// TIA Portal project "N16-1166-5_27082020" (V13) (continued)

               #IFM_Switch_State := #IFM_Switch_State + 1;
           1:
               // set number of pulses to send to the IFM senzor
               #IFM_Pulse_Number := #IFM_ApplicationIndex;
               //change the state to the next value
               #IFM_Switch_State := #IFM_Switch_State + 1;
           2:
               //pulsing in precisely time intervals
               IF #IFM_Pulse_Number > 0 THEN
                   IF #IFM_Input_2 = false AND #IFM_Timer_State = 0 THEN
                       #IFM_Input_2 := true;
                       #IFM_Timer_State := #IFM_Pulse_Period / 2;
                   ELSIF #IFM_Input_2 = true AND #IFM_Timer_State = 0 THEN
                       #IFM_Input_2 := false;
                       #IFM_Timer_State := #IFM_Pulse_Period / 2;
                       #IFM_Pulse_Number := #IFM_Pulse_Number - 1;
                   END_IF;
               ELSE
                   #IFM_Switch_State := #IFM_Switch_State + 1;
               END_IF;
           3:
               // set input 1 to false
               #IFM_Input_1 := false;
               //set to init state
               #IFM_Switch_State := 0;
               //set free to switch of application       
               #IFM_PulsApplicationSwitch := true;
           ELSE  // Statement section ELSE
               #IFM_Switch_State := 0;
               #IFM_Input_1 := false;
               #IFM_Input_2 := false;
       END_CASE;
   ELSE
       #IFM_PulsApplicationSwitch := false;
   END_IF;
   *)
END_FUNCTION_BLOCK

FUNCTION_BLOCK "vacuum_cleaner_controll"   // FB2, SCL
{ S7_Optimized_Access := 'FALSE' }
VERSION : 0.1
BEGIN

   IF #vacuum_sensor = true THEN
       #switch := true;
       #timer_lib_Instance.lock := false;
       #vacuum_control_variable := true;
   END_IF;

   IF #switch = true THEN
       #timer_lib_Instance(time_value := #vacuum_cleaner_activity_interval);
       IF #timer_lib_Instance.DONE = true THEN
           #switch := false;
           #vacuum_control_variable := false;
       END_IF;
   END_IF;
END_FUNCTION_BLOCK

FUNCTION_BLOCK "RPA30_F_TRIGR"   // FB4, SCL
{ S7_Optimized_Access := 'FALSE' }
VERSION : 0.1
BEGIN

   IF #PREVIOS = true AND #CLK = false THEN
       #Q := true;
       #STATE := true;
   ELSE
       #Q := false;
   END_IF;

   #PREVIOS := #CLK;
END_FUNCTION_BLOCK

FUNCTION_BLOCK "PA30_IFM_point_checking"   // FB5, SCL
{ S7_Optimized_Access := 'FALSE' }
VERSION : 0.1
BEGIN




   IF #execute = true THEN
   (*
   ** if keyence are disabled in its checking
   *)
       IF #checking_state >= 30 AND #keyence_enable = false THEN
           #checking_state := 27;
       END_IF;

       #index := 0;
       #mark := 0;
       #temp_string := '';

       //pars input data from left ifm sensor 
       WHILE #index < "RPA30_DataBlock".pa30_right_size_in DO
           IF "RPA30_DataBlock".pa30_left_ifm_data[#index] = '#' THEN
               IF #mark > 1 THEN
                   #left_camera_points_pixel[#mark - 1] := STRING_TO_UINT(#temp_string);
                   #temp_string := '';
               END_IF;

               #mark := #mark + 1;
           ELSE
               IF #mark > 1 THEN
                   #temp_string := CONCAT(IN1 := #temp_string, IN2 := "RPA30_DataBlock".pa30_left_ifm_data[#index]);
               END_IF;
           END_IF;

           #index := #index + 1;
       END_WHILE;

       #index := 0;
       #mark := 0;
       #temp_string := '';

       //pars input data from right ifm sensor
       WHILE #index < "RPA30_DataBlock".pa30_right_size_in DO
           IF "RPA30_DataBlock".pa30_right_ifm_data[#index] = '#' THEN
               IF #mark > 1 THEN
                   #right_camera_points_pixel[#mark - 1] := STRING_TO_UINT(#temp_string);
                   #temp_string := '';
               END_IF;

               #mark := #mark + 1;
           ELSE
               IF #mark > 1 THEN
                   #temp_string := CONCAT(IN1 := #temp_string, IN2 := "RPA30_DataBlock".pa30_right_ifm_data[#index]);
               END_IF;
           END_IF;

           #index := #index + 1;
       END_WHILE;

       IF #ifm_side > 0 THEN
           CASE #checking_state OF
               0, 1:  // nastavení senzorů
                   #DONE := false;
                   #checking_state := 2;

               2:
   (* kontrola zda byla aplikace přepnuta *)
                   IF 1 = "RPA30_DataBlock".pa30_left_ifm_actived_application_index AND
                       1 = "RPA30_DataBlock".pa30_right_ifm_actived_application_index THEN
                       #checking_state := 3;
                   END_IF;

               3:
   (* čekání na deaktivaci senzoru *)
                   IF #left_camera_points_pixel[((#ifm_side - 1) * 2) + 1] = 0 THEN
                       #checking_state := 4;
                   END_IF;

               4:
   (* čekání na aktivaci senzoru na bodě L1 a následné přepnutí kamery na bod L2*)
                   IF #left_camera_points_pixel[((#ifm_side - 1) * 2) + 1] > #pixel_treshold THEN
                       #checking_state := 5;
                       #beep := true;
                       #points := 1;
                   END_IF;

               5:
   (* čekání na deaktivaci senzoru *)
                   IF (#left_camera_points_pixel[((#ifm_side - 1) * 2) + 1] = #left_camera_points_pixel[((#ifm_side - 1) * 2) + 2]) = 0 THEN
                       #checking_state := 6;
                   END_IF;

               6:
   (* čekání na aktivaci senzoru  *)
                   IF #left_camera_points_pixel[((#ifm_side - 1) * 2) + 2] > #pixel_treshold THEN
                       #checking_state := 7;
                       #beep := true;
                       #points := 2;
                   END_IF;
               7:
   (* čekání na deaktivaci obou senzorů *)
                   IF (#left_camera_points_pixel[((#ifm_side - 1) * 2) + 2] + #right_camera_points_pixel[((#ifm_side - 1) * 3) + 1]) = 0 THEN
                       #checking_state := 8;
                   END_IF;

               8:
   (* čekání na aktivaci obou senzorů a následné přepnutí senzoru na bod P2 *)
                   IF #right_camera_points_pixel[((#ifm_side - 1) * 3) + 1] > #pixel_treshold THEN
                       #beep := true;
                       #points := 3;
                       #checking_state := 9;
                   END_IF;
               9:
                   IF (#right_camera_points_pixel[((#ifm_side - 1) * 3) + 1] + #right_camera_points_pixel[((#ifm_side - 1) * 3) + 2]) = 0 THEN
                       #checking_state := 10;
                   END_IF;
               10:
                   IF #right_camera_points_pixel[((#ifm_side - 1) * 3) + 2] > #pixel_treshold THEN
                       #beep := true;
                       #points := 4;
                       #checking_state := 11;
                   END_IF;

               11:
                   IF (#right_camera_points_pixel[((#ifm_side - 1) * 3) + 2] + #right_camera_points_pixel[((#ifm_side - 1) * 3) + 3]) = 0 THEN
                       #checking_state := 12;
                   END_IF;
               12:
                   IF #right_camera_points_pixel[((#ifm_side - 1) * 3) + 3] > #pixel_treshold THEN
                       #beep := true;
                       #points := 5;

                       IF #ifm_side = 2 OR "RPA30_DataBlock".RPA30_station_configuration = 0 THEN
                           #checking_state := 27;
                       ELSE
                           IF #keyence_enable = true THEN
                               #checking_state := 30;
                           ELSE
                               #checking_state := 27;
                           END_IF;
                       END_IF;
                   END_IF;
               30:
                   //sensor 1 non active
                   IF (#ifm_side = 1 AND "RPA30_keyence_left_1" = false) OR (#ifm_side = 3 AND "RPA30_keyence_left_2" = false) THEN
                       #checking_state := 31;
                   END_IF;
               31:
                   //sensor 1 active
                   IF (#ifm_side = 1 AND "RPA30_keyence_left_1" = true) OR #ifm_side = 3 AND "RPA30_keyence_left_2" = true THEN
                       #checking_state := 32;
                       #points := 6;
                       #beep := true;
                   END_IF;
               32:
                   //sensor 1 non active
                   IF (#ifm_side = 1 AND "RPA30_keyence_left_1" = false) OR (#ifm_side = 3 AND "RPA30_keyence_left_2" = false) THEN
                       #checking_state := 33;
                   END_IF;

               33:
                   //sensor 2 non active
                   IF (#ifm_side = 1 AND "RPA30_keyence_middle_2" = false) OR (#ifm_side = 3 AND "RPA30_keyence_middle_1" = false) THEN
                       #checking_state := 34;
                   END_IF;

               34:
                   //sensor 2 active
                   IF (#ifm_side = 1 AND "RPA30_keyence_middle_2" = true) OR #ifm_side = 3 AND ("RPA30_keyence_middle_1" = true) THEN
                       #checking_state := 35;
                       #points := 7;
                       #beep := true;
                   END_IF;
               35:
                   //sensor 2 non active
                   IF (#ifm_side = 1 AND "RPA30_keyence_middle_2" = false) OR (#ifm_side = 3 AND "RPA30_keyence_middle_1" = false) THEN
                       #checking_state := 36;
                   END_IF;
               36:
                   //sensor 3 non active
                   IF (#ifm_side = 1 AND "RPA30_keyence_right_1" = false) OR (#ifm_side = 3 AND "RPA30_keyence_right_2" = false) THEN
                       #checking_state := 37;
                   END_IF;
               37:
                   //sensor 3 atvite
                   IF (#ifm_side = 1 AND "RPA30_keyence_right_1" = true) OR (#ifm_side = 3 AND "RPA30_keyence_right_2" = true) THEN
                       #checking_state := 27;
                       #points := 8;
                       #beep := true;
                   END_IF;
               27:
                   #DONE := true;
          END_CASE;
      END_IF;
   ELSE
       #checking_state := 0;
       #points := 0;
       #DONE := false;
   END_IF;

   (* pípnutí při zachycení bodu *)
   IF #beep = true THEN
       #timer_lib_Instance(100);
       IF #timer_lib_Instance.DONE = false THEN
           #primerbox_siren := true;
       ELSE
           #primerbox_siren := false;
           #beep := false;
       END_IF;
   END_IF;
END_FUNCTION_BLOCK

FUNCTION_BLOCK "O2VxEth1500"   // FB8, SCL
TITLE = O2VxEth1500 for S7-15xx CPU FW V1.7 or higher
{ S7_Optimized_Access := 'FALSE' }
AUTHOR : ifm-sytl
FAMILY : O2Vx
NAME : O2Vx1500
VERSION : 1.3
// Basic Application program for O2Vx
// connected to S7-1500 station via CPU-internal Ethernet interface
// for S7-15xx CPU Firmware V1.7 or higher
BEGIN
END_FUNCTION_BLOCK

FUNCTION_BLOCK "fs_scaner_fce"   // FB11, SCL
{ S7_Optimized_Access := 'FALSE' }
VERSION : 0.1
BEGIN
   #Receive_P2P_Instance(BUFFER:=#Receive_P2P_Instance.ReceiveBuffer,"PORT" := "FS~CM_PtP_1");

   IF #Receive_P2P_Instance.NDR = true THEN
      Chars_TO_Strg(Chars:=#Receive_P2P_Instance.ReceiveBuffer,
                    pChars:=0,
                    Cnt:=#Receive_P2P_Instance.received_length-1,
                    Strg=>#scaner_input_data);
   END_IF;
END_FUNCTION_BLOCK

FUNCTION_BLOCK "print_label_PA60"   // FB13, SCL
{ S7_Optimized_Access := 'FALSE' }
VERSION : 0.1
BEGIN

   #DONE := false;

   IF #TCON_Instance.DONE = false THEN
       #TCON_Instance.REQ := NOT #TCON_Instance.REQ;
       #TCON_Instance(CONNECT := "printer_connection",
                               ID := 10);
   ELSE
       //date formating
       #date_string := CONCAT(IN1 := #date_string, IN2 := "copyAndFill"(characterFill := '0', charReplace := '+', stringIn := (DELETE(IN := INT_TO_STRING(#"date".DAY), L := 1, P := 1)), P := 0, char_number := 2));
       #date_string := CONCAT(IN1 := #date_string, IN2 := '.');
       #date_string := CONCAT(IN1 := #date_string, IN2 := "copyAndFill"(characterFill := '0', charReplace := '+', stringIn := (DELETE(IN := INT_TO_STRING(#"date".MONTH), L := 1, P := 1)), P := 0, char_number := 2));
       #date_string := CONCAT(IN1 := #date_string, IN2 := '.');
       #date_string := CONCAT(IN1 := #date_string, IN2 := "copyAndFill"(characterFill := '0', charReplace := '+', stringIn := (DELETE(IN := UINT_TO_STRING(#"date".YEAR), L := 1, P := 1)), P := 0, char_number := 4));

       //time formating
       #time_string := CONCAT(IN1 := #time_string, IN2 := "copyAndFill"(characterFill := '0', charReplace := '+', stringIn := (DELETE(IN := INT_TO_STRING(#"date".HOUR), L := 1, P := 1)), P := 0, char_number := 2));
       #time_string := CONCAT(IN1 := #time_string, IN2 := ':');
       #time_string := CONCAT(IN1 := #time_string, IN2 := "copyAndFill"(characterFill := '0', charReplace := '+', stringIn := (DELETE(IN := INT_TO_STRING(#"date".MINUTE), L := 1, P := 1)), P := 0, char_number := 2));
       #time_string := CONCAT(IN1 := #time_string, IN2 := ':');
       #time_string := CONCAT(IN1 := #time_string, IN2 := "copyAndFill"(characterFill := '0', charReplace := '+', stringIn := (DELETE(IN := INT_TO_STRING(#"date".SECOND), L := 1, P := 1)), P := 0, char_number := 2));

       //qr code string formating
       IF #frame_conf = 0 THEN
           #MCode := 'AU581*1762975*';
       ELSE
           #MCode := 'AU326-1*1768362*';
       END_IF;

       #MCode := CONCAT(IN1 := #MCode, IN2 := #date_string);
       #MCode := CONCAT(IN1 := #MCode, IN2 := '*');
       #MCode := CONCAT(IN1 := #MCode, IN2 := #time_string);
       #MCode := CONCAT(IN1 := #MCode, IN2 := '*172');
       #MCode := CONCAT(IN1 := #MCode, IN2 := #order);

       //send command to the printer
       IF #TSEND_Instance.DONE = false THEN

       #numberOfChar := 0;
       Strg_TO_Chars(Strg := '^XA^MMT^PW480^LL0200^LS0^FO0,0^GFA,03072,03072,00032,:Z64:eJztk7GO4jAQhifJIZ2gIYWbrbZchTdI5Ui3PUjx+1jQ8RRZaCK7uTI3vNz9M4YEpIu47nQSI+wYO1/GM/MP0cte9k/NbXW2c+ehm+Y/8nb8StaOu5m7raKSG5mLMJ3Hv+WT56rHlE88jcvEm1mevcz1IP554nl88QkflF/O+X/GZ1H5VU8V4s/TZh7G+K8v',
                     pChars := #chars,
                     Cnt => #chars,
                     Chars := #data_out);

       #numberOfChar := #numberOfChar +#chars;
       Strg_TO_Chars(Strg := 'mi0+lLXGUoYvGSfb7sF/HvALPS1D8CEc5V9/zy9cmznXknPGOvfp2kWqbIr/bXhjzi/MVDN75iMPWFz5THjj4NQ58K5RHhvJPzzCfxXCPqhvecI/Nrzy39S/s8Kl0RJ4pzzix4vdqo9+c4jneIgxHgIV8R0L5W1ZlmvwZBp4b3CLzxbbGZaSWvUalj3ucApU7dNA/oOvurv8C9+SAYvLK09GjvgofP2Lmc+IXsaBO7pAATV4eIT/0uxw3V3ic',
                     pChars := #numberOfChar,
                     Cnt => #chars,
                     Chars := #data_out);

       #numberOfChar := #numberOfChar + #chars;
       Strg_TO_Chars(Strg := 'Q+kEsVUPpyEr3pMJ2Qfo/KSBohhqfwPSYB75CWMKx+V33wh3HNPGxk+xq+IZlgpvyspW4NX/ShvzR0vNac+dEH1V0kOfC5/sVA+9W8z8cjIHV8PeOuDOxQ7R8gnDE/1T77Fb0S0Jao35d8S0oH8aWqvneeR7n24agCeVQj+xi/Ap/qLhhqQt/rTSjqlQPWj1t5HfXax32j9adEmFT7qz476085LKoT+EbTewav+5GSR4qeb/o2T/J',
                     pChars := #numberOfChar,
                     Cnt => #chars,
                     Chars := #data_out);

       #numberOfChar := #numberOfChar + #chars;
       Strg_TO_Chars(Strg := 'PoX9sxH7QLEPxQMA9UX1B/aYOC9SRTXhQnjWfxPfTPVsJKysolSYRLVLjtEkt5YHT0PTWwTfysKf8xf678ev5c7f3J+cte9rL/zn4DEoMnnA==:C58E',
                     pChars := #numberOfChar,
                     Cnt => #chars,
                     Chars := #data_out);

       #numberOfChar := #numberOfChar + #chars;
       IF #frame_conf = 0 THEN
           Strg_TO_Chars(Strg := '^FT32,85^A0N,17,16^FH\^FDAU581^FS^FT32,104^A0N,17,16^FH\^FDID-No. 1762975^FS^FT180,122^A0N,17,16^FH\^FD',
                         pChars := #numberOfChar,
                         Cnt => #chars,
                         Chars := #data_out);
       ELSE //zde upravit kód rámu
           Strg_TO_Chars(Strg := '^FT32,85^A0N,17,16^FH\^FDAU326-1^FS^FT32,104^A0N,17,16^FH\^FDID-No. 1768362^FS^FT180,122^A0N,17,16^FH\^FD',
                         pChars := #numberOfChar,
                         Cnt => #chars,
                         Chars := #data_out);
       END_IF;

       #numberOfChar := #numberOfChar + #chars;
       Strg_TO_Chars(Strg := #time_string,
                     pChars := #numberOfChar,
                     Cnt => #chars,
                     Chars := #data_out);

       #numberOfChar := #numberOfChar + #chars;
       Strg_TO_Chars(Strg := '^FS^FT31,142^A0N,17,16^FH\^FDSerial-No:^FS',
                         pChars := #numberOfChar,
                         Cnt => #chars,
                         Chars := #data_out);

       #numberOfChar := #numberOfChar + #chars;
       Strg_TO_Chars(Strg := '^BY96,96^FT332,141^BXN,4,200,0,0,1,~^FH\^FD',
                     pChars := #numberOfChar,
                     Cnt => #chars,
                     Chars := #data_out);

       #numberOfChar := #numberOfChar + #chars;
       Strg_TO_Chars(Strg := #MCode,
                     pChars := #numberOfChar,
                     Cnt => #chars,
                     Chars := #data_out);

       #numberOfChar := #numberOfChar + #chars;
       Strg_TO_Chars(Strg := '^FS^FT32,161^A0N,17,16^FH\^FDWBR Made in Romania (WRO)^FS^FT31,123^A0N,17,16^FH\^FDDate:^FS^FT31,181^A0N,17,16^FH\^FD',
                     pChars := #numberOfChar,
                     Cnt => #chars,
                     Chars := #data_out);

       #numberOfChar := #numberOfChar + #chars;
       Strg_TO_Chars(Strg := #MCode,
                     pChars := #numberOfChar,
                     Cnt => #chars,
                     Chars := #data_out);

       #numberOfChar := #numberOfChar + #chars;
       Strg_TO_Chars(Strg := '^FS^FT70,122^A0N,17,16^FH\^FD',
                     pChars := #numberOfChar,
                     Cnt => #chars,
                     Chars := #data_out);

       #numberOfChar := #numberOfChar + #chars;
       Strg_TO_Chars(Strg := #date_string,
                     pChars := #numberOfChar,
                     Cnt => #chars,
                     Chars := #data_out);

       #numberOfChar := #numberOfChar + #chars;
       Strg_TO_Chars(Strg := '^FS^FT179,142^A0N,17,16^FH\^FD',
                     pChars := #numberOfChar,
                     Cnt => #chars,
                     Chars := #data_out);

       #numberOfChar := #numberOfChar + #chars;
       Strg_TO_Chars(Strg := #order,
                     pChars := #numberOfChar,
                     Cnt => #chars,
                     Chars := #data_out);

       #numberOfChar := #numberOfChar + #chars;
       Strg_TO_Chars(Strg := '^FS^FT114,142^A0N,17,16^FH\^FD172^FS^PQ1,0,1,Y^XZ',
                     pChars := #numberOfChar,
                     Cnt => #chars,
                     Chars := #data_out);

       #numberOfChar := #numberOfChar + #chars;


           #TSEND_Instance.REQ := NOT #TSEND_Instance.REQ;
           #TSEND_Instance(ID := 10,LEN := #numberOfChar, DATA := #data_out);
       ELSE
           IF #TDISCON_Instance.DONE = false THEN
               #TDISCON_Instance.REQ := NOT #TDISCON_Instance.REQ;
               #TDISCON_Instance(ID := 10);
           ELSE
               #TDISCON_Instance.DONE := false;
               #TSEND_Instance.DONE := false;
               #TCON_Instance.DONE := false;
               #DONE := true;
           END_IF;
       END_IF;
   END_IF;
END_FUNCTION_BLOCK

FUNCTION_BLOCK "bottle_changing"   // FB14, SCL
{ S7_Optimized_Access := 'FALSE' }
VERSION : 0.1
BEGIN

   #DONE := false;

   CASE #"step" OF
      0:  // take secound bottle than will used
          IF #bottle = 1 THEN
              #hmi_label_index := 28;
              #use_bottle_2 := true ;
              #use_bottle_1 := false;
          ELSIF #bottle = 2 THEN
              #hmi_label_index := 29;
              #use_bottle_2 := false;
              #use_bottle_1 := true;
          END_IF;



          IF (#bottle_presence_sensor_1 = false AND  #bottle = 2) OR (#bottle_presence_sensor_2 = false AND  #bottle = 1) THEN
              #"step" := 10;
              #take_bottle := true;
          END_IF;

      10: // scan label and check expiration
          #hmi_label_index := "RPA10B_hmi_scan_bottle";
          IF "RPA10B_Scanner_DB".NDR = true THEN
              IF RD_SYS_T(#current_time) < 0 THEN
                  ;
              END_IF;

              #bottle_checking_result := "bottle_label_check"(input_data := "RPA10B_datablock".RPA10B_scanned_data, chemical_type := 5);

              IF #bottle_checking_result = 0 THEN
                  IF  #bottle_presence_sensor_2 = false  THEN
                      #bottle_label_2 := "RPA10B_datablock".RPA10B_scanned_data;
                  ELSIF #bottle_presence_sensor_1 = false THEN
                      #bottle_label_1 := "RPA10B_datablock".RPA10B_scanned_data;
                  END_IF;

                  IF (#bottle = 1 AND #bottle_presence_sensor_2 = false) OR (#bottle = 2 AND #bottle_presence_sensor_2 = false) THEN
                      #"step" := 40;
                  ELSIF (#bottle = 1 AND #bottle_presence_sensor_1 = false) OR (#bottle = 2 AND #bottle_presence_sensor_1 = false) THEN
                      #"step" := 20;
                  END_IF;

              ELSIF #bottle_checking_result = 2 THEN
                  "RPA10B_datablock".PA10B_error_state_lock := 400;
                  #"step" := 30;
              ELSIF #bottle_checking_result = 3 THEN
                  "RPA10B_datablock".PA10B_error_state_lock := 401;
                  #"step" := 30;
              ELSIF #bottle_checking_result = 4 THEN
                  "RPA10B_datablock".PA10B_error_state_lock := 402;
                  #"step" := 30;
              ELSIF #bottle_checking_result = 5 THEN
                  "RPA10B_datablock".PA10B_error_state_lock := 403;
                  #"step" := 30;
              END_IF;
          END_IF;

      20: //change pad bottle 1
          #hmi_label_index := "RPA10B_hmi_change_pad";
          "RPA10B_datablock".RPA10B_show_pad_left := true;
          IF "RPA10B_change_pad"(padSensor := "RPA10B_primerbox_pad_sensor_left",
                                     padIsChangedButton := "RPA10B_primerbox_button_PAD_IS_CHANGED",
                                     failStatelockIdetifier := 6,
                                     bigFailStateLock := "RPA10B_datablock".PA10B_big_fail_state_lock,
                                     FatalErrorStateLock := "RPA10B_datablock".PA10B_fatal_error_state_lock,
                                     readyLED => "RPA10B_primerbox_LED_green_ready",
                                     notReadyLED => "RPA10B_primerbox_LED_red_NOT_READY",
                                     changePedLED => "RPA10B_primerbox_LED_orange_change_pad",
                                     confirmButtonLED => "RPA10B_LCD_LED_blue_confirm_button",
                                     failStateLock := "RPA10B_datablock".PA10B_fail_state_lock) THEN
              "RPA10B_datablock".RPA10B_show_pad_left := false;
              #bottle_1_cyclus_counter := 0;
              IF RD_SYS_T(#bottle_1_expiration) < 2 THEN
                  IF (#bottle = 2 AND #bottle_presence_sensor_1 = false) OR (#bottle = 1 AND #bottle_presence_sensor_2 = false) THEN
                      #"step" := 50;
                  ELSE
                      #"step" := 60;
                  END_IF;
              END_IF;
          END_IF;

      30: // bottle expired
          IF "RPA10B_datablock".PA10B_error_state_lock = 400 OR "RPA10B_datablock".PA10B_error_state_lock = 401 OR "RPA10B_datablock".PA10B_error_state_lock = 402 OR "RPA10B_datablock".PA10B_error_state_lock = 403 THEN
              "RPA10B_LCD_LED_blue_confirm_button" := "Clock_0.5Hz";
              IF "RPA10B_LCD_button_confirm" = true THEN
                  "RPA10B_datablock".PA10B_error_state_lock := 0;
                  "RPA10B_LCD_LED_blue_confirm_button" := false;
                  #"step" := 10;
              END_IF;
          END_IF;

      40: // change pad bottle 2
          #hmi_label_index := "RPA10B_hmi_change_pad";
          "RPA10B_datablock".RPA10B_show_pad_right := true;
          IF "RPA10B_change_pad"(padSensor := "RPA10B_primerbox_pad_sensor_right",
                                     padIsChangedButton := "RPA10B_primerbox_button_PAD_IS_CHANGED",
                                     failStatelockIdetifier := 6,
                                     bigFailStateLock := "RPA10B_datablock".PA10B_big_fail_state_lock,
                                     FatalErrorStateLock := "RPA10B_datablock".PA10B_fatal_error_state_lock,
                                     readyLED => "RPA10B_primerbox_LED_green_ready",
                                     notReadyLED => "RPA10B_primerbox_LED_red_NOT_READY",
                                     changePedLED => "RPA10B_primerbox_LED_orange_change_pad",
                                     confirmButtonLED => "RPA10B_LCD_LED_blue_confirm_button",
                                     failStateLock := "RPA10B_datablock".PA10B_fail_state_lock) THEN
              "RPA10B_datablock".RPA10B_show_pad_right := false;
              #bottle_2_cyclus_counter := 0;
              IF RD_SYS_T(#bottle_2_expiration) < 2 THEN
                  IF (#bottle = 1 AND #bottle_presence_sensor_2 = false) OR (#bottle = 2 AND #bottle_presence_sensor_1 = false) THEN
                      #"step" := 50;
                  ELSE
                      #"step" := 60;
                  END_IF;
              END_IF;
          END_IF;

      50: // put bottle back to primerbox and take secound bottle
          IF #bottle_presence_sensor_1 = true AND #bottle_presence_sensor_2 = true THEN
              #take_bottle := false;
              IF #bottle = 1 THEN
                  //choose bottle 1
                  #hmi_label_index := 28;
                  #use_bottle_2 := false;
                  #use_bottle_1 := true;
              ELSIF #bottle = 2 THEN
                  //choose bottle 2
                  #hmi_label_index := 29;
                  #use_bottle_2 := true;
                  #use_bottle_1 := false;
              END_IF;
          ELSE
              //put bottle back to primer box
              #hmi_label_index := 30;
          END_IF;

          IF (#bottle = 1 AND #bottle_presence_sensor_1 = false) OR (#bottle = 2 AND #bottle_presence_sensor_2 = false) THEN
              #take_bottle := true;
              #"step" := 10;
          END_IF;

      60: //end
          #DONE := true;
          #"step" := 0;
       ELSE  // Statement section ELSE
           #"step" := 0;
   END_CASE;
END_FUNCTION_BLOCK

FUNCTION_BLOCK "fs_print_label_fce"   // FB15, SCL
{ S7_Optimized_Access := 'FALSE' }
VERSION : 0.1
BEGIN
END_FUNCTION_BLOCK

FUNCTION_BLOCK "shaker_door_lock_control"   // FB18, SCL
{ S7_Optimized_Access := 'FALSE' }
VERSION : 0.1
BEGIN


   #mixer_1_door_1_lock := #mixer_1_presence_sensor_1 AND #mixer_1_door_1_is_close AND #mixer_door_lock_enable[0];
   #mixer_1_door_2_lock := #mixer_1_presence_sensor_2 AND #mixer_1_door_2_is_close AND #mixer_door_lock_enable[1];
   #mixer_2_door_1_lock := #mixer_2_presence_sensor_1 AND #mixer_2_door_1_is_close AND #mixer_door_lock_enable[2];
   #mixer_2_door_2_lock := #mixer_2_presence_sensor_2 AND #mixer_2_door_2_is_close AND #mixer_door_lock_enable[3];
   #mixer_3_door_1_lock := (#mixer_3_presence_sensor_1 AND #mixer_3_door_1_is_close AND #mixer_door_lock_enable[4]);
END_FUNCTION_BLOCK

FUNCTION_BLOCK "print_label_582"   // FB19, SCL
{ S7_Optimized_Access := 'FALSE' }
VERSION : 0.1
BEGIN





   #DONE := false;

   IF #TCON_Instance.DONE = false THEN
       #TCON_Instance.REQ := NOT #TCON_Instance.REQ;
       #TCON_Instance(CONNECT := "printer_connection",
                               ID := 10);
   ELSE

       //date formating
       #date_string := CONCAT(IN1 := #date_string, IN2 := "copyAndFill"(characterFill := '0', charReplace := '+', stringIn := (DELETE(IN := INT_TO_STRING(#"date".DAY), L := 1, P := 1)), P := 0, char_number := 2));
       #date_string := CONCAT(IN1 := #date_string, IN2 := '.');
       #date_string := CONCAT(IN1 := #date_string, IN2 := "copyAndFill"(characterFill := '0', charReplace := '+', stringIn := (DELETE(IN := INT_TO_STRING(#"date".MONTH), L := 1, P := 1)), P := 0, char_number := 2));
       #date_string := CONCAT(IN1 := #date_string, IN2 := '.');
       #date_string := CONCAT(IN1 := #date_string, IN2 := "copyAndFill"(characterFill := '0', charReplace := '+', stringIn := (DELETE(IN := UINT_TO_STRING(#"date".YEAR), L := 1, P := 1)), P := 0, char_number := 4));

       //time formating
       #time_string := CONCAT(IN1 := #time_string, IN2 := "copyAndFill"(characterFill := '0', charReplace := '+', stringIn := (DELETE(IN := INT_TO_STRING(#"date".HOUR), L := 1, P := 1)), P := 0, char_number := 2));
       #time_string := CONCAT(IN1 := #time_string, IN2 := ':');
       #time_string := CONCAT(IN1 := #time_string, IN2 := "copyAndFill"(characterFill := '0', charReplace := '+', stringIn := (DELETE(IN := INT_TO_STRING(#"date".MINUTE), L := 1, P := 1)), P := 0, char_number := 2));
       #time_string := CONCAT(IN1 := #time_string, IN2 := ':');
       #time_string := CONCAT(IN1 := #time_string, IN2 := "copyAndFill"(characterFill := '0', charReplace := '+', stringIn := (DELETE(IN := INT_TO_STRING(#"date".SECOND), L := 1, P := 1)), P := 0, char_number := 2));

       //qr code string formating
       #MCode := 'AU582*1762976*';
       #MCode := CONCAT(IN1 := #MCode, IN2 := #date_string);
       #MCode := CONCAT(IN1 := #MCode, IN2 := '*');
       #MCode := CONCAT(IN1 := #MCode, IN2 := #time_string);
       #MCode := CONCAT(IN1 := #MCode, IN2 := '*172');
       #MCode := CONCAT(IN1 := #MCode, IN2 := #order_string);

       //command formating
       #command := CONCAT(IN1 := #command, IN2 := '^XA');
       #command := CONCAT(IN1 := #command, IN2 := #label1);
       //...next data in the label

       //barcode
       #command := CONCAT(IN1 := #command, IN2 := '^BY96,96^FT270,145^BXN,4,200,0,0,1,~^FH\^FD');
       #command := CONCAT(IN1 := #command, IN2 := #MCode);
       #command := CONCAT(IN1 := #command, IN2 := '^FS');

       //label
       #command := CONCAT(IN1 := #command, IN2 := '^FT31,181^A0N,16,14^FH\^FD');
       #command := CONCAT(IN1 := #command, IN2 := #MCode);
       #command := CONCAT(IN1 := #command, IN2 := '^FS');

       //date
       #command := CONCAT(IN1 := #command, IN2 := '^FT70,122^A0N,17,16^FH\^FD');
       #command := CONCAT(IN1 := #command, IN2 := #date_string);
       #command := CONCAT(IN1 := #command, IN2 := '^FS');
       Strg_TO_Chars(Strg := #command,
                     pChars := 0,
                     Cnt => #chars,
                     Chars := #data_out);

       #command := '';
       //time
       #command := CONCAT(IN1 := #command, IN2 := '^FT180,122^A0N,17,16^FH\^FD');
       #command := CONCAT(IN1 := #command, IN2 := #time_string);
       #command := CONCAT(IN1 := #command, IN2 := '^FS');

       //order part 1
       #command := CONCAT(IN1 := #command, IN2 := '^FT114,142^A0N,17,16^FH\^FD172^FS');

       //#order part 2
       #command := CONCAT(IN1 := #command, IN2 := '^FT179,142^A0N,17,16^FH\^FD');
       #command := CONCAT(IN1 := #command, IN2 := #order_string);
       #command := CONCAT(IN1 := #command, IN2 := '^FS');

       #command := CONCAT(IN1 := #command, IN2 := '^XZ');

       //prepeare to send

       #numberOfChar := #chars;
       Strg_TO_Chars(Strg := #command,
                     pChars := #chars,
                     Cnt => #chars,
                     Chars := #data_out);

       #numberOfChar := #numberOfChar + #chars;

       //send command to the printer
       IF #TSEND_Instance.DONE = false THEN
           #TSEND_Instance.REQ := NOT #TSEND_Instance.REQ;
           #TSEND_Instance(ID := 1,LEN := #numberOfChar, DATA := #data_out);
       ELSE
           IF #TDISCON_Instance.DONE = false THEN
               #TDISCON_Instance.REQ := NOT #TDISCON_Instance.REQ;
               #TDISCON_Instance(ID := 1);
           ELSE
               #TDISCON_Instance.DONE := false;
               #TSEND_Instance.DONE := false;
               #TCON_Instance.DONE := false;
               #DONE := true;
           END_IF;
       END_IF;
   END_IF;
END_FUNCTION_BLOCK

FUNCTION_BLOCK "scaner_runtime"   // FB20, SCL
{ S7_Optimized_Access := 'FALSE' }
VERSION : 0.1
BEGIN
   #fs_scaner_fce_Instance();


   IF #fs_scaner_fce_Instance.Receive_P2P_Instance.NDR = true THEN
       IF #shaker_index = 0 THEN
           IF #filling_e = false AND #print_sp_bottle_e = false AND #chemical_type > 0 THEN
               IF #fs_scaner_fce_Instance.scaner_input_data[LEN(#fs_scaner_fce_Instance.scaner_input_data)] = 'M' THEN
                   #filling_e := true;
               ELSE
                   #print_sp_bottle_e := true;
               END_IF;
           END_IF;
       END_IF;
   END_IF;
END_FUNCTION_BLOCK

FUNCTION_BLOCK "timer_lib"   // FB21, SCL
{ S7_Optimized_Access := 'FALSE' }
VERSION : 0.1
BEGIN
   #DONE := false;
   IF #lock = true THEN
       IF RD_LOC_T(#actual_time) < 2 THEN
           IF TIME_TO_DINT(IN := T_DIFF(IN1 := #actual_time, IN2 := #"time")) > #time_value THEN
               #DONE := true;
               #lock := false;
           END_IF;
       END_IF;
   ELSE
       IF RD_LOC_T(#"time") < 2 THEN
           #lock := true;
       END_IF;
   END_IF;
END_FUNCTION_BLOCK

FUNCTION_BLOCK "filling_station_main"   // FB23, SCL
{ S7_Optimized_Access := 'FALSE' }
VERSION : 0.1
BEGIN

   IF #fs_activity_state = true THEN
       (* station internal state runtime control *)
       "fs_internal_state"(switch_automat_manual := "ib_FS_LCD_switch_automat_manual",
                           tcp_connection := "tcp_datablock".tcp_connection,
                           confirm_button := "ib_FS_LCD_button_confirm",
                           error_state := #fs_error_state,
                           confirm_led := "ob_FS_LCD_confirm_button_LED_blue",
                           beacon_green := "ob_FS_LCD_beacon_green",
                           beacon_orange := "ob_FS_LCD_beacon_orange",
                           beacon_red := "ob_FS_LCD_beacon_red",
                           beacon_siren := "ob_FS_LCD_beacon_siren",
                           alarm:=#fs_alarm);

       IF #fs_reset_enable = true THEN
           "station_reset"(funel_1:="ob_FS_move_UP_funel_1",
                           funel_2:="ob_FS_move_UP_funel_2",
                           funel_3:="ob_FS_move_UP_funel_3",
                           funel_4:="ob_FS_move_UP_funel_4",
                           funel_5:="ob_FS_move_UP_funel_5",
                           fs_reset_e:=#fs_reset_enable,
                           fs_chemical_type:=#chemical_type,
                           fill_bottle_step:=#fce_filling_Instance."step",
                           shake_deinit:=#sp_bottle_shaking_Instance.shake_deinit,
                           print_sp_bottle_label_step:=#fce_print_sp_botle_label_Instance."step",
                           fs_show_manual_or_scan:=#manual_or_scan,
                           fs_show_button:=#fs_show_button,
                           fs_show_fill_button:=#fce_filling_Instance.show_fill_button,
                           fs_funel_control:=#fce_filling_Instance.funel_control,
                           hmi_label_index:=#hmi_label_index);
       END_IF;

       IF #filling_enable = false AND #print_sp_bottle_label_enable = false AND #shaking_enable = false THEN
           IF #chemical_type > 0 AND #chemical_type < 3 THEN
               #hmi_label_index := 21;
               #fs_show_button := true;
               #manual_or_scan := false;
           ELSIF #chemical_type > 2 THEN
               IF #chemical_type_pre = 0 AND #chemical_type > 2 THEN
                   #manual_or_scan := true;
               END_IF;

               IF #manual_or_scan = false THEN
                   #hmi_label_index := 22;
               ELSE
                   #hmi_label_index := 20;
               END_IF;

               #fs_show_button := true;
           ELSIF #chemical_type = 0 THEN
               #fs_show_button := false;
               #manual_or_scan := false;
               #hmi_label_index := 0;
           END_IF;
       ELSE
           #fs_show_button := true;
           #manual_or_scan := false;
       END_IF;

       #chemical_type_pre := #chemical_type;

       (* scanner runtime hadler and input data parsing *)
       #scaner_runtime_Instance(shaker_index:=#sp_bottle_shaking_Instance.runtime_shaker_index_finding_Instance.shaker_index,
                                chemical_type:=#chemical_type,
                                filling_e:=#filling_enable,
                                print_sp_bottle_e:=#print_sp_bottle_label_enable);

       (* print suplier bottle label work cycle *)
       IF #shaking_enable = false THEN // shaking work cycle is more important
           #fce_print_sp_botle_label_Instance(scanned_data := #scaner_runtime_Instance.fs_scaner_fce_Instance.scaner_input_data,
                                              scaner_ndr := #scaner_runtime_Instance.fs_scaner_fce_Instance.Receive_P2P_Instance.NDR,
                                              expire_time_Primer_DV954V1 := #expire_time_Primer_DV954V1,
                                              expire_time_Activator_DW646 := #expire_time_Activator_DW646,
                                              expire_time_Remover_SIKA_208 := #expire_time_Remover_SIKA_208,
                                              expire_time_Primer_SIKA_207 := #expire_time_Primer_SIKA_207,
                                              expire_time_Activator_SIKA_110 := #expire_time_Activator_SIKA_110,
                                              print_sp_bottle_label_enable := #print_sp_bottle_label_enable,
                                              error_state := #fs_error_state,
                                              fs_SIKA_remover_order := #fs_SIKA_remover_order,
                                              fs_SIKA_primer_order := #fs_SIKA_primer_order,
                                              fs_SIKA_activator_order := #fs_SIKA_activator_order,
                                              shake_enable := #shaking_enable,
                                              chemical_type := #chemical_type,
                                              show_button := #fs_show_button,
                                              hmi_label_index := #hmi_label_index,
                                              show_manual_input := #manual_or_scan);

           (*small bottle filling work cycle*)

           #fce_filling_Instance(scanned_data := #scaner_runtime_Instance.fs_scaner_fce_Instance.scaner_input_data,
                                 scaner_ndr := #scaner_runtime_Instance.fs_scaner_fce_Instance.Receive_P2P_Instance.NDR,
                                 funel_1_bottle_presence := "ib_FS_sensor_bottle_1",
                                 funel_2_bottle_presence := "ib_FS_sensor_bottle_2",
                                 funel_3_bottle_presence := "ib_FS_sensor_bottle_3",
                                 funel_4_bottle_presence := "ib_FS_sensor_bottle_4",
                                 funel_5_bottle_presence := "ib_FS_sensor_bottle_5",
                                 primer_DV954V1_time_after_shaking := #primer_DV954V1_time_after_shaking,
                                 primer_SIKA_207_time_after_shaking := #primer_SIKA_207_time_after_shaking,
                                 filling_enable := #filling_enable,
                                 chemical_type := #chemical_type,
                                 shaking_enable := #shaking_enable,
                                 error_state := #fs_error_state,
                                 move_UP_funel_1 := "ob_FS_move_UP_funel_1",
                                 move_UP_funel_2 := "ob_FS_move_UP_funel_2",
                                 move_UP_funel_3 := "ob_FS_move_UP_funel_3",
                                 move_UP_funel_4 := "ob_FS_move_UP_funel_4",
                                 move_UP_funel_5 := "ob_FS_move_UP_funel_5",
                                 hmi_label_index := #hmi_label_index);

       END_IF;

       (* shaking fce *)


       #sp_bottle_shaking_Instance(shaker_1_door_1_lock := "ob_FS_mixer_1_door_1_lock",
                                   shaker_1_door_2_lock := "ob_FS_mixer_1_door_2_lock",
                                   shaker_2_door_1_lock := "ob_FS_mixer_2_door_1_lock",
                                   shaker_2_door_2_lock := "ob_FS_mixer_2_door_2_lock",
                                   shaker_3_door_1_lock := "ob_FS_mixer_3_door_lock",
                                   chemical_type := #chemical_type,
                                   error_state := #fs_error_state,
                                   shaker_1_door_1_bottle_presence := "ib_FS_mixer_1_presence_sensor_1",
                                   shaker_1_door_2_bottle_presence := "ib_FS_mixer_1_presence_sensor_2",
                                   shaker_2_door_1_bottle_presence := "ib_FS_mixer_2_presence_sensor_1",
                                   shaker_2_door_2_bottle_presence := "ib_FS_mixer_2_presence_sensor_2",
                                   shaker_3_door_1_bottle_presence := "ib_FS_mixer_3_bottle_pressence",
                                   shaker_1_door_1_position := "ib_FS_mixer_1_door_1_is_close",
                                   shaker_1_door_2_position := "ib_FS_mixer_1_door_2_is_close",
                                   shaker_2_door_1_position := "ib_FS_mixer_2_door_1_is_close",
                                   shaker_2_door_2_position := "ib_FS_mixer_2_door_2_is_close",
                                   shaker_3_door_1_position := "ib_FS_mixer_3_door_position",
                                   shaking_enable := #shaking_enable,
                                   scaner_ndr := #scaner_runtime_Instance.fs_scaner_fce_Instance.Receive_P2P_Instance.NDR,
                                   scanned_data := #scaner_runtime_Instance.fs_scaner_fce_Instance.scaner_input_data,
                                   hmi_label_index := #hmi_label_index);


   ELSE
       (* inactive station state *)
       "station_inactive_state"(fs_start_button:="ib_FS_LCD_button_start",
                                fune_1:="ob_FS_move_UP_funel_1",
                                fune_2:="ob_FS_move_UP_funel_2",
                                fune_3:="ob_FS_move_UP_funel_3",
                                fune_4:="ob_FS_move_UP_funel_4",
                                fune_5:="ob_FS_move_UP_funel_5",
                                fs_reset_enable:=#fs_reset_enable,
                                fs_start_led:="ob_FS_LCD_start_button_LED_green",
                                error_state:=#fs_error_state,
                                beacon_red:="ob_FS_LCD_beacon_red",
                                beacon_orange:="ob_FS_LCD_beacon_orange",
                                beacon_green:="ob_FS_LCD_beacon_green",
                                beacon_siren:="ob_FS_LCD_beacon_siren",
                                fs_station_activity:=#fs_activity_state,
                                chemical_type:=#chemical_type,
                                fill_bottle_step:=#fce_filling_Instance."step",
                                shake_deinit:=#sp_bottle_shaking_Instance.shake_deinit,
                                print_sp_bottle_label_step:=#fce_print_sp_botle_label_Instance."step",
                                fs_show_manual_or_scan:=#manual_or_scan,
                                fs_show_button:=#fs_show_button,
                                fs_show_fill_button:=#fce_filling_Instance.show_fill_button,
                                fs_funel_control:=#fce_filling_Instance.funel_control,
                                hmi_label_index:=#hmi_label_index);
   END_IF;
END_FUNCTION_BLOCK

FUNCTION_BLOCK "sp_bottle_shaking"   // FB24, SCL
{ S7_Optimized_Access := 'FALSE' }
VERSION : 0.1
BEGIN
   (* runtime checking shaker state *)
   #runtime_shaker_index_finding_Instance(mixer_1_presence_sensor_1:=#shaker_1_door_1_bottle_presence,
                                          mixer_1_presence_sensor_2:=#shaker_1_door_2_bottle_presence,
                                          mixer_2_presence_sensor_1:=#shaker_2_door_1_bottle_presence,
                                          mixer_2_presence_sensor_2:=#shaker_2_door_2_bottle_presence,
                                          mixer_3_presence_sensor_1:=#shaker_3_door_1_bottle_presence,
                                          error_state_identifier:=#error_state,
                                          shaking_enable:=#shaking_enable);
   (* shaking work cycle *)
   IF #shaking_enable = true THEN
       IF #runtime_shaker_index_finding_Instance.shaker_index = 1 THEN
           IF #shaker_1_door_1_position THEN
               #hmi_label_index := 5;
               IF #scaner_ndr = true THEN
                   #label_scanned := true;
               END_IF;

               IF #shaker_1_door_1_lock THEN
                   IF RD_SYS_T(#runtime_shake_count_expiration_Instance.fs_mixer_expiration[#runtime_shaker_index_finding_Instance.shaker_index - 1]) < 2 THEN
                       ;
                   END_IF;
                   #shake_deinit := true;
               END_IF;
           ELSE
               #hmi_label_index := 15;
           END_IF;
       ELSIF #runtime_shaker_index_finding_Instance.shaker_index = 2 THEN
           IF #shaker_1_door_2_position THEN
               #hmi_label_index := 5;
               IF #scaner_ndr = true THEN
                   #label_scanned := true;
               END_IF;

               IF #shaker_1_door_2_lock THEN
                   IF RD_SYS_T(#runtime_shake_count_expiration_Instance.fs_mixer_expiration[#runtime_shaker_index_finding_Instance.shaker_index - 1]) < 2 THEN
                       ;
                   END_IF;
                   #shake_deinit := true;
               END_IF;
           ELSE
               #hmi_label_index := 15;
           END_IF;
       ELSIF #runtime_shaker_index_finding_Instance.shaker_index = 3 THEN
           IF #shaker_2_door_1_position THEN
               #hmi_label_index := 5;
               IF #scaner_ndr = true THEN
                   #label_scanned := true;
               END_IF;

               IF #shaker_2_door_1_lock THEN
                   IF RD_SYS_T(#runtime_shake_count_expiration_Instance.fs_mixer_expiration[#runtime_shaker_index_finding_Instance.shaker_index - 1]) < 2 THEN
                       ;
                   END_IF;
                   #shake_deinit := true;
               END_IF;
           ELSE
               #hmi_label_index := 15;
           END_IF;
       ELSIF #runtime_shaker_index_finding_Instance.shaker_index = 4 THEN
           IF #shaker_2_door_2_position THEN
               #hmi_label_index := 5;
               IF #scaner_ndr = true THEN
                   #label_scanned := true;
               END_IF;

               IF #shaker_2_door_2_lock THEN
                   IF RD_SYS_T(#runtime_shake_count_expiration_Instance.fs_mixer_expiration[#runtime_shaker_index_finding_Instance.shaker_index - 1]) < 2 THEN
                       ;
                   END_IF;
                   #shake_deinit := true;
               END_IF;
           ELSE
               #hmi_label_index := 15;
           END_IF;
       ELSIF #runtime_shaker_index_finding_Instance.shaker_index = 5 THEN
           IF #shaker_3_door_1_position THEN
               #hmi_label_index := 5;
               IF #scaner_ndr = true THEN
                   #label_scanned := true;
               END_IF;

               IF #shaker_3_door_1_lock THEN
                   IF RD_SYS_T(#runtime_shake_count_expiration_Instance.fs_mixer_expiration[#runtime_shaker_index_finding_Instance.shaker_index - 1]) < 2 THEN
                       ;
                   END_IF;
                   #shake_deinit := true;
               END_IF;
           ELSE
               #hmi_label_index := 15;
           END_IF;
       ELSIF #runtime_shaker_index_finding_Instance.shaker_index = 0 THEN
           #hmi_label_index := 3;

           (* check shaker state befor start shaking procedur and wait for inserting bottle inside shaker and set up shaker index *)
           IF (#chemical_type = 4 AND #shaker_3_door_1_bottle_presence = true) OR
               ((#chemical_type < 4 OR #chemical_type = 5) AND
               #shaker_1_door_1_bottle_presence AND
               #shaker_1_door_2_bottle_presence AND
               #shaker_2_door_1_bottle_presence AND
               #shaker_2_door_2_bottle_presence) THEN
               (* no free shaker *)
               #shake_deinit := true;
               #error_state := 512;
           END_IF;
       END_IF;

       IF #label_scanned THEN
           "parse_scanned_label"(scanned_data:=#scanned_data,
                                 chemical:=#chemical,
                                 batch_no:=#batch_no,
                                 expire_date_time:=#expire_date_time,
                                 filling_opening_date_time:=#filling_opening_date_time,
                                 bottle_type:=#bottle_type);

           IF #bottle_type = 'M' THEN
               #database_command_done := "get_table_record_item"(table := 'suplier_bottle',
                                                                 record := #batch_no,
                                                                 item := 'last_shake',
                                                                 record_key := 'batch_code',
                                                                 server_connection := "tcp_datablock".tcp_connection,
                                                                 index := "tcp_datablock".fs_fill_bottle_index,
                                                                 output_buffer := #temp_buffer);
               IF #database_command_done = true THEN

                   #input_string := "parse_input_data"(#temp_buffer);
                   IF #input_string <> 'ERROR' THEN
                       IF RD_SYS_T(#current_time) < 2 THEN
                           ;
                       END_IF;

